REGION Network 343
   RUNG wire#powerrail
      Contact( "EMS".Carrier[46].SDC_OUT.Faults.CarrierSpacingFault )
      Coil( "Carrier_46_Carrier_Spacing_Fault" )
   END_RUNG
   // the same network as SCL:
   "Carrier_46_Carrier_Spacing_Fault" := "EMS".Carrier[46].SDC_OUT.Faults.CarrierSpacingFault;
END_REGION

REGION Network 344
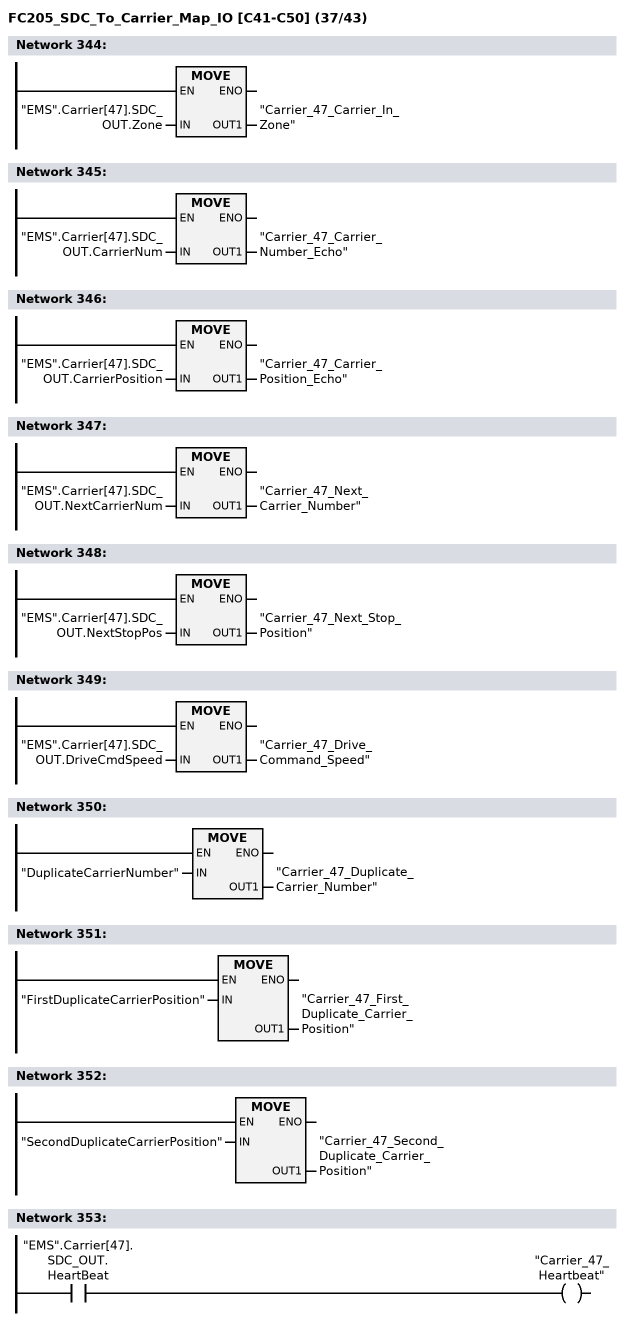
   RUNG wire#powerrail
      Move(in := "EMS".Carrier[47].SDC_OUT.Zone, out1 => "Carrier_47_Carrier_In_Zone")
   END_RUNG
   // the same network as SCL:
   "Carrier_47_Carrier_In_Zone" := "EMS".Carrier[47].SDC_OUT.Zone;
END_REGION

REGION Network 345
   RUNG wire#powerrail
      Move(in := "EMS".Carrier[47].SDC_OUT.CarrierNum, out1 => "Carrier_47_Carrier_Number_Echo")
   END_RUNG
   // the same network as SCL:
   "Carrier_47_Carrier_Number_Echo" := "EMS".Carrier[47].SDC_OUT.CarrierNum;
END_REGION

REGION Network 346
   RUNG wire#powerrail
      Move(in := "EMS".Carrier[47].SDC_OUT.CarrierPosition, out1 => "Carrier_47_Carrier_Position_Echo")
   END_RUNG
   // the same network as SCL:
   "Carrier_47_Carrier_Position_Echo" := "EMS".Carrier[47].SDC_OUT.CarrierPosition;
END_REGION

REGION Network 347
   RUNG wire#powerrail
      Move(in := "EMS".Carrier[47].SDC_OUT.NextCarrierNum, out1 => "Carrier_47_Next_Carrier_Number")
   END_RUNG
   // the same network as SCL:
   "Carrier_47_Next_Carrier_Number" := "EMS".Carrier[47].SDC_OUT.NextCarrierNum;
END_REGION

REGION Network 348
   RUNG wire#powerrail
      Move(in := "EMS".Carrier[47].SDC_OUT.NextStopPos, out1 => "Carrier_47_Next_Stop_Position")
   END_RUNG
   // the same network as SCL:
   "Carrier_47_Next_Stop_Position" := "EMS".Carrier[47].SDC_OUT.NextStopPos;
END_REGION

REGION Network 349
   RUNG wire#powerrail
      Move(in := "EMS".Carrier[47].SDC_OUT.DriveCmdSpeed, out1 => "Carrier_47_Drive_Command_Speed")
   END_RUNG
   // the same network as SCL:
   "Carrier_47_Drive_Command_Speed" := "EMS".Carrier[47].SDC_OUT.DriveCmdSpeed;
END_REGION

REGION Network 350
   RUNG wire#powerrail
      Move(in := "DuplicateCarrierNumber", out1 => "Carrier_47_Duplicate_Carrier_Number")
   END_RUNG
   // the same network as SCL:
   "Carrier_47_Duplicate_Carrier_Number" := "DuplicateCarrierNumber";
END_REGION

REGION Network 351
   RUNG wire#powerrail
      Move(in := "FirstDuplicateCarrierPosition", out1 => "Carrier_47_First_Duplicate_Carrier_Position")
   END_RUNG
   // the same network as SCL:
   "Carrier_47_First_Duplicate_Carrier_Position" := "FirstDuplicateCarrierPosition";
END_REGION

REGION Network 352
   RUNG wire#powerrail
      Move(in := "SecondDuplicateCarrierPosition", out1 => "Carrier_47_Second_Duplicate_Carrier_Position")
   END_RUNG
   // the same network as SCL:
   "Carrier_47_Second_Duplicate_Carrier_Position" := "SecondDuplicateCarrierPosition";
END_REGION

REGION Network 353
   RUNG wire#powerrail
      Contact( "EMS".Carrier[47].SDC_OUT.HeartBeat )
      Coil( "Carrier_47_Heartbeat" )
   END_RUNG
   // the same network as SCL:
   "Carrier_47_Heartbeat" := "EMS".Carrier[47].SDC_OUT.HeartBeat;
END_REGION

REGION Network 354
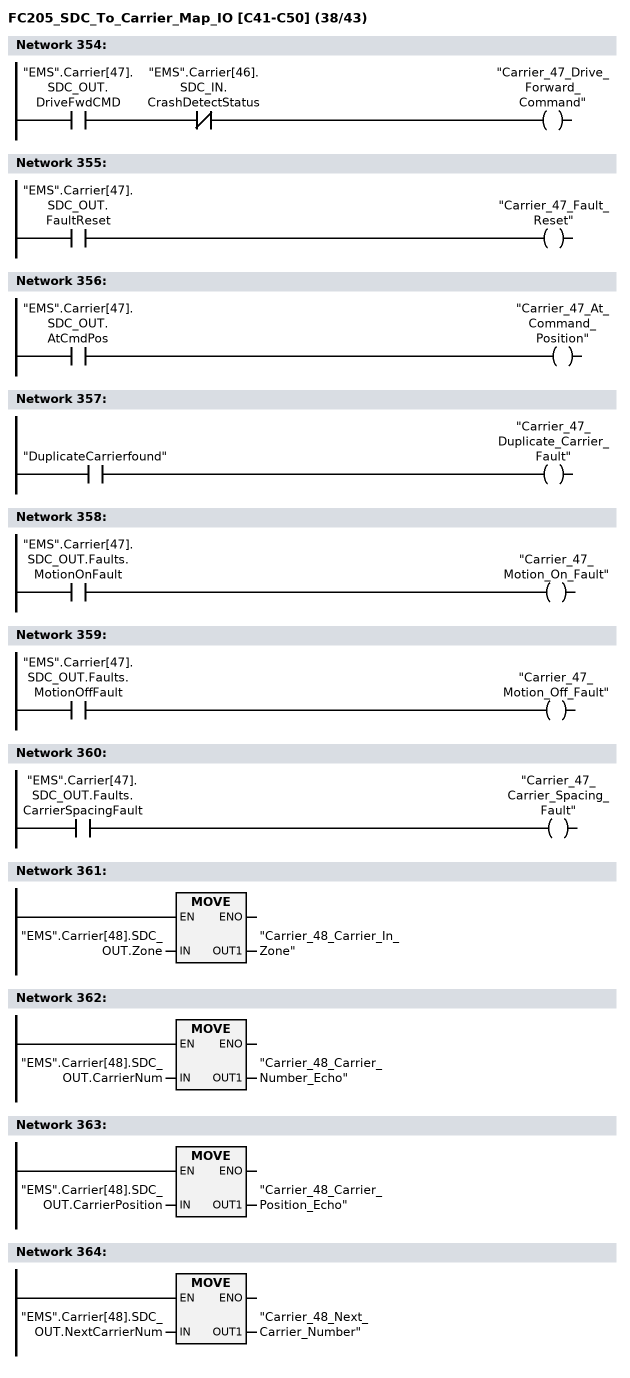
   RUNG wire#powerrail
      Contact( "EMS".Carrier[47].SDC_OUT.DriveFwdCMD )
      I_Contact( "EMS".Carrier[46].SDC_IN.CrashDetectStatus )
      Coil( "Carrier_47_Drive_Forward_Command" )
   END_RUNG
   // the same network as SCL:
   "Carrier_47_Drive_Forward_Command" := "EMS".Carrier[47].SDC_OUT.DriveFwdCMD AND NOT "EMS".Carrier[46].SDC_IN.CrashDetectStatus;
END_REGION

REGION Network 355
   RUNG wire#powerrail
      Contact( "EMS".Carrier[47].SDC_OUT.FaultReset )
      Coil( "Carrier_47_Fault_Reset" )
   END_RUNG
   // the same network as SCL:
   "Carrier_47_Fault_Reset" := "EMS".Carrier[47].SDC_OUT.FaultReset;
END_REGION

REGION Network 356
   RUNG wire#powerrail
      Contact( "EMS".Carrier[47].SDC_OUT.AtCmdPos )
      Coil( "Carrier_47_At_Command_Position" )
   END_RUNG
   // the same network as SCL:
   "Carrier_47_At_Command_Position" := "EMS".Carrier[47].SDC_OUT.AtCmdPos;
END_REGION

REGION Network 357
   RUNG wire#powerrail
      Contact( "DuplicateCarrierfound" )
      Coil( "Carrier_47_Duplicate_Carrier_Fault" )
   END_RUNG
   // the same network as SCL:
   "Carrier_47_Duplicate_Carrier_Fault" := "DuplicateCarrierfound";
END_REGION

REGION Network 358
   RUNG wire#powerrail
      Contact( "EMS".Carrier[47].SDC_OUT.Faults.MotionOnFault )
      Coil( "Carrier_47_Motion_On_Fault" )
   END_RUNG
   // the same network as SCL:
   "Carrier_47_Motion_On_Fault" := "EMS".Carrier[47].SDC_OUT.Faults.MotionOnFault;
END_REGION

REGION Network 359
   RUNG wire#powerrail
      Contact( "EMS".Carrier[47].SDC_OUT.Faults.MotionOffFault )
      Coil( "Carrier_47_Motion_Off_Fault" )
   END_RUNG
   // the same network as SCL:
   "Carrier_47_Motion_Off_Fault" := "EMS".Carrier[47].SDC_OUT.Faults.MotionOffFault;
END_REGION

REGION Network 360
   RUNG wire#powerrail
      Contact( "EMS".Carrier[47].SDC_OUT.Faults.CarrierSpacingFault )
      Coil( "Carrier_47_Carrier_Spacing_Fault" )
   END_RUNG
   // the same network as SCL:
   "Carrier_47_Carrier_Spacing_Fault" := "EMS".Carrier[47].SDC_OUT.Faults.CarrierSpacingFault;
END_REGION

REGION Network 361
   RUNG wire#powerrail
      Move(in := "EMS".Carrier[48].SDC_OUT.Zone, out1 => "Carrier_48_Carrier_In_Zone")
   END_RUNG
   // the same network as SCL:
   "Carrier_48_Carrier_In_Zone" := "EMS".Carrier[48].SDC_OUT.Zone;
END_REGION

REGION Network 362
   RUNG wire#powerrail
      Move(in := "EMS".Carrier[48].SDC_OUT.CarrierNum, out1 => "Carrier_48_Carrier_Number_Echo")
   END_RUNG
   // the same network as SCL:
   "Carrier_48_Carrier_Number_Echo" := "EMS".Carrier[48].SDC_OUT.CarrierNum;
END_REGION

REGION Network 363
   RUNG wire#powerrail
      Move(in := "EMS".Carrier[48].SDC_OUT.CarrierPosition, out1 => "Carrier_48_Carrier_Position_Echo")
   END_RUNG
   // the same network as SCL:
   "Carrier_48_Carrier_Position_Echo" := "EMS".Carrier[48].SDC_OUT.CarrierPosition;
END_REGION

REGION Network 364
   RUNG wire#powerrail
      Move(in := "EMS".Carrier[48].SDC_OUT.NextCarrierNum, out1 => "Carrier_48_Next_Carrier_Number")
   END_RUNG
   // the same network as SCL:
   "Carrier_48_Next_Carrier_Number" := "EMS".Carrier[48].SDC_OUT.NextCarrierNum;
END_REGION

REGION Network 365
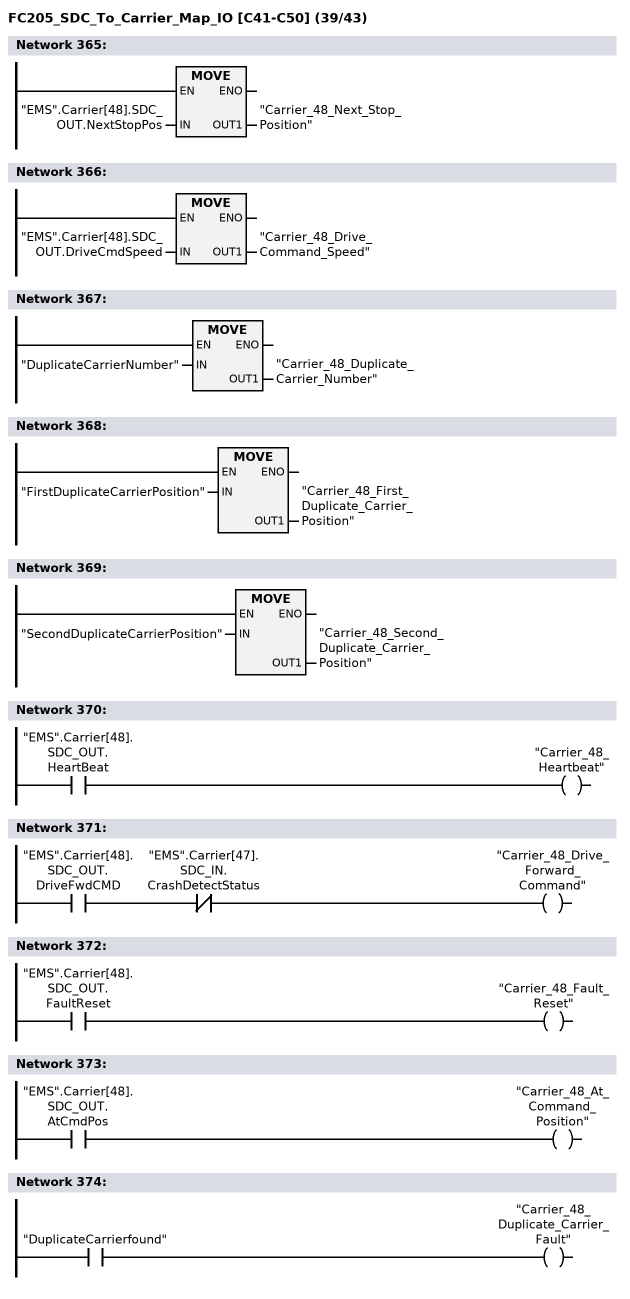
   RUNG wire#powerrail
      Move(in := "EMS".Carrier[48].SDC_OUT.NextStopPos, out1 => "Carrier_48_Next_Stop_Position")
   END_RUNG
   // the same network as SCL:
   "Carrier_48_Next_Stop_Position" := "EMS".Carrier[48].SDC_OUT.NextStopPos;
END_REGION

REGION Network 366
   RUNG wire#powerrail
      Move(in := "EMS".Carrier[48].SDC_OUT.DriveCmdSpeed, out1 => "Carrier_48_Drive_Command_Speed")
   END_RUNG
   // the same network as SCL:
   "Carrier_48_Drive_Command_Speed" := "EMS".Carrier[48].SDC_OUT.DriveCmdSpeed;
END_REGION

REGION Network 367
   RUNG wire#powerrail
      Move(in := "DuplicateCarrierNumber", out1 => "Carrier_48_Duplicate_Carrier_Number")
   END_RUNG
   // the same network as SCL:
   "Carrier_48_Duplicate_Carrier_Number" := "DuplicateCarrierNumber";
END_REGION

REGION Network 368
   RUNG wire#powerrail
      Move(in := "FirstDuplicateCarrierPosition", out1 => "Carrier_48_First_Duplicate_Carrier_Position")
   END_RUNG
   // the same network as SCL:
   "Carrier_48_First_Duplicate_Carrier_Position" := "FirstDuplicateCarrierPosition";
END_REGION

REGION Network 369
   RUNG wire#powerrail
      Move(in := "SecondDuplicateCarrierPosition", out1 => "Carrier_48_Second_Duplicate_Carrier_Position")
   END_RUNG
   // the same network as SCL:
   "Carrier_48_Second_Duplicate_Carrier_Position" := "SecondDuplicateCarrierPosition";
END_REGION

REGION Network 370
   RUNG wire#powerrail
      Contact( "EMS".Carrier[48].SDC_OUT.HeartBeat )
      Coil( "Carrier_48_Heartbeat" )
   END_RUNG
   // the same network as SCL:
   "Carrier_48_Heartbeat" := "EMS".Carrier[48].SDC_OUT.HeartBeat;
END_REGION

REGION Network 371
   RUNG wire#powerrail
      Contact( "EMS".Carrier[48].SDC_OUT.DriveFwdCMD )
      I_Contact( "EMS".Carrier[47].SDC_IN.CrashDetectStatus )
      Coil( "Carrier_48_Drive_Forward_Command" )
   END_RUNG
   // the same network as SCL:
   "Carrier_48_Drive_Forward_Command" := "EMS".Carrier[48].SDC_OUT.DriveFwdCMD AND NOT "EMS".Carrier[47].SDC_IN.CrashDetectStatus;
END_REGION

REGION Network 372
   RUNG wire#powerrail
      Contact( "EMS".Carrier[48].SDC_OUT.FaultReset )
      Coil( "Carrier_48_Fault_Reset" )
   END_RUNG
   // the same network as SCL:
   "Carrier_48_Fault_Reset" := "EMS".Carrier[48].SDC_OUT.FaultReset;
END_REGION

REGION Network 373
   RUNG wire#powerrail
      Contact( "EMS".Carrier[48].SDC_OUT.AtCmdPos )
      Coil( "Carrier_48_At_Command_Position" )
   END_RUNG
   // the same network as SCL:
   "Carrier_48_At_Command_Position" := "EMS".Carrier[48].SDC_OUT.AtCmdPos;
END_REGION

REGION Network 374
   RUNG wire#powerrail
      Contact( "DuplicateCarrierfound" )
      Coil( "Carrier_48_Duplicate_Carrier_Fault" )
   END_RUNG
   // the same network as SCL:
   "Carrier_48_Duplicate_Carrier_Fault" := "DuplicateCarrierfound";
END_REGION

REGION Network 375
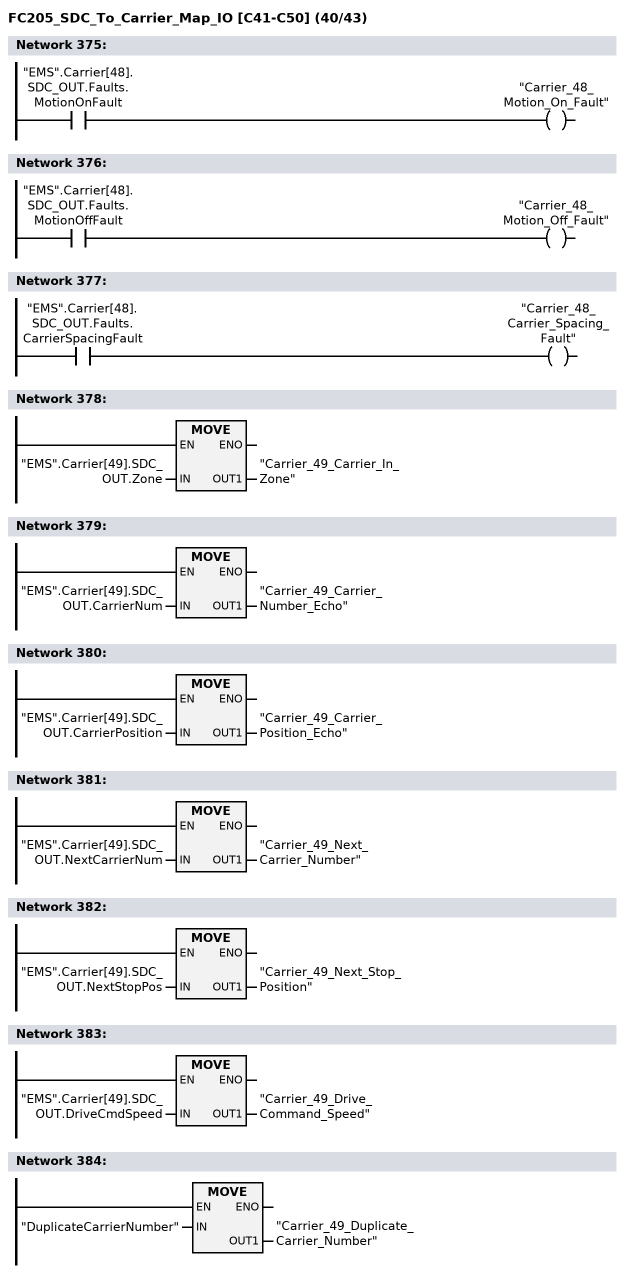
   RUNG wire#powerrail
      Contact( "EMS".Carrier[48].SDC_OUT.Faults.MotionOnFault )
      Coil( "Carrier_48_Motion_On_Fault" )
   END_RUNG
   // the same network as SCL:
   "Carrier_48_Motion_On_Fault" := "EMS".Carrier[48].SDC_OUT.Faults.MotionOnFault;
END_REGION

REGION Network 376
   RUNG wire#powerrail
      Contact( "EMS".Carrier[48].SDC_OUT.Faults.MotionOffFault )
      Coil( "Carrier_48_Motion_Off_Fault" )
   END_RUNG
   // the same network as SCL:
   "Carrier_48_Motion_Off_Fault" := "EMS".Carrier[48].SDC_OUT.Faults.MotionOffFault;
END_REGION

REGION Network 377
   RUNG wire#powerrail
      Contact( "EMS".Carrier[48].SDC_OUT.Faults.CarrierSpacingFault )
      Coil( "Carrier_48_Carrier_Spacing_Fault" )
   END_RUNG
   // the same network as SCL:
   "Carrier_48_Carrier_Spacing_Fault" := "EMS".Carrier[48].SDC_OUT.Faults.CarrierSpacingFault;
END_REGION

REGION Network 378
   RUNG wire#powerrail
      Move(in := "EMS".Carrier[49].SDC_OUT.Zone, out1 => "Carrier_49_Carrier_In_Zone")
   END_RUNG
   // the same network as SCL:
   "Carrier_49_Carrier_In_Zone" := "EMS".Carrier[49].SDC_OUT.Zone;
END_REGION

REGION Network 379
   RUNG wire#powerrail
      Move(in := "EMS".Carrier[49].SDC_OUT.CarrierNum, out1 => "Carrier_49_Carrier_Number_Echo")
   END_RUNG
   // the same network as SCL:
   "Carrier_49_Carrier_Number_Echo" := "EMS".Carrier[49].SDC_OUT.CarrierNum;
END_REGION

REGION Network 380
   RUNG wire#powerrail
      Move(in := "EMS".Carrier[49].SDC_OUT.CarrierPosition, out1 => "Carrier_49_Carrier_Position_Echo")
   END_RUNG
   // the same network as SCL:
   "Carrier_49_Carrier_Position_Echo" := "EMS".Carrier[49].SDC_OUT.CarrierPosition;
END_REGION

REGION Network 381
   RUNG wire#powerrail
      Move(in := "EMS".Carrier[49].SDC_OUT.NextCarrierNum, out1 => "Carrier_49_Next_Carrier_Number")
   END_RUNG
   // the same network as SCL:
   "Carrier_49_Next_Carrier_Number" := "EMS".Carrier[49].SDC_OUT.NextCarrierNum;
END_REGION

REGION Network 382
   RUNG wire#powerrail
      Move(in := "EMS".Carrier[49].SDC_OUT.NextStopPos, out1 => "Carrier_49_Next_Stop_Position")
   END_RUNG
   // the same network as SCL:
   "Carrier_49_Next_Stop_Position" := "EMS".Carrier[49].SDC_OUT.NextStopPos;
END_REGION

REGION Network 383
   RUNG wire#powerrail
      Move(in := "EMS".Carrier[49].SDC_OUT.DriveCmdSpeed, out1 => "Carrier_49_Drive_Command_Speed")
   END_RUNG
   // the same network as SCL:
   "Carrier_49_Drive_Command_Speed" := "EMS".Carrier[49].SDC_OUT.DriveCmdSpeed;
END_REGION

REGION Network 384
   RUNG wire#powerrail
      Move(in := "DuplicateCarrierNumber", out1 => "Carrier_49_Duplicate_Carrier_Number")
   END_RUNG
   // the same network as SCL:
   "Carrier_49_Duplicate_Carrier_Number" := "DuplicateCarrierNumber";
END_REGION

REGION Network 385
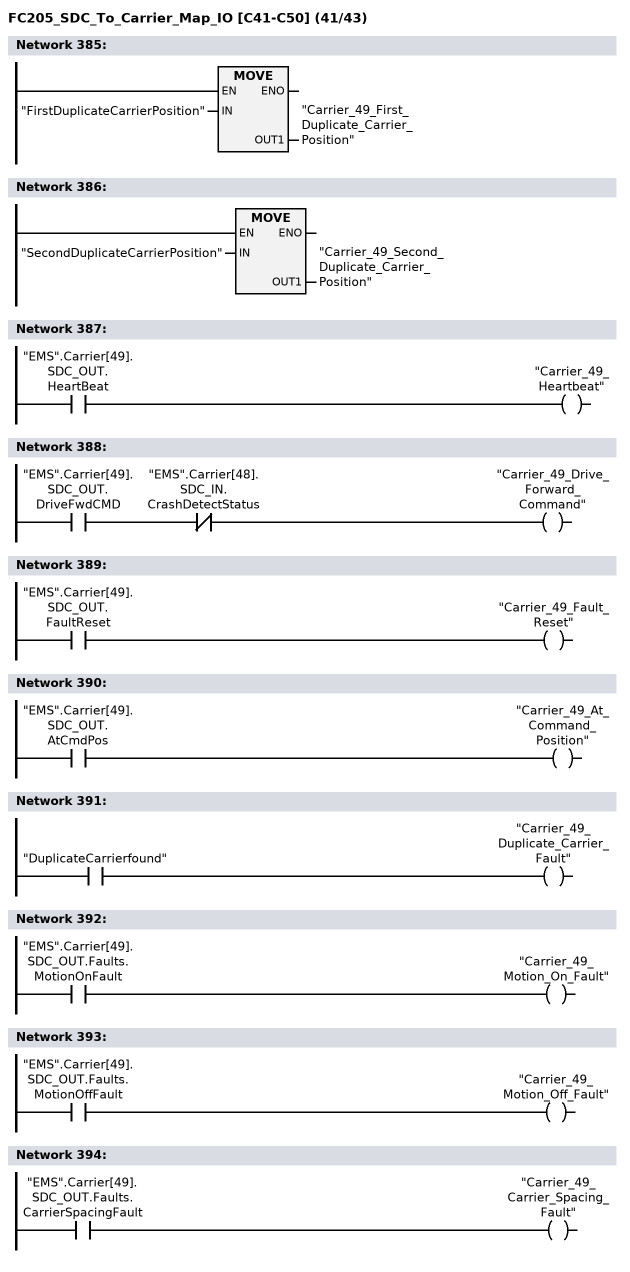
   RUNG wire#powerrail
      Move(in := "FirstDuplicateCarrierPosition", out1 => "Carrier_49_First_Duplicate_Carrier_Position")
   END_RUNG
   // the same network as SCL:
   "Carrier_49_First_Duplicate_Carrier_Position" := "FirstDuplicateCarrierPosition";
END_REGION

REGION Network 386
   RUNG wire#powerrail
      Move(in := "SecondDuplicateCarrierPosition", out1 => "Carrier_49_Second_Duplicate_Carrier_Position")
   END_RUNG
   // the same network as SCL:
   "Carrier_49_Second_Duplicate_Carrier_Position" := "SecondDuplicateCarrierPosition";
END_REGION

REGION Network 387
   RUNG wire#powerrail
      Contact( "EMS".Carrier[49].SDC_OUT.HeartBeat )
      Coil( "Carrier_49_Heartbeat" )
   END_RUNG
   // the same network as SCL:
   "Carrier_49_Heartbeat" := "EMS".Carrier[49].SDC_OUT.HeartBeat;
END_REGION

REGION Network 388
   RUNG wire#powerrail
      Contact( "EMS".Carrier[49].SDC_OUT.DriveFwdCMD )
      I_Contact( "EMS".Carrier[48].SDC_IN.CrashDetectStatus )
      Coil( "Carrier_49_Drive_Forward_Command" )
   END_RUNG
   // the same network as SCL:
   "Carrier_49_Drive_Forward_Command" := "EMS".Carrier[49].SDC_OUT.DriveFwdCMD AND NOT "EMS".Carrier[48].SDC_IN.CrashDetectStatus;
END_REGION

REGION Network 389
   RUNG wire#powerrail
      Contact( "EMS".Carrier[49].SDC_OUT.FaultReset )
      Coil( "Carrier_49_Fault_Reset" )
   END_RUNG
   // the same network as SCL:
   "Carrier_49_Fault_Reset" := "EMS".Carrier[49].SDC_OUT.FaultReset;
END_REGION

REGION Network 390
   RUNG wire#powerrail
      Contact( "EMS".Carrier[49].SDC_OUT.AtCmdPos )
      Coil( "Carrier_49_At_Command_Position" )
   END_RUNG
   // the same network as SCL:
   "Carrier_49_At_Command_Position" := "EMS".Carrier[49].SDC_OUT.AtCmdPos;
END_REGION

REGION Network 391
   RUNG wire#powerrail
      Contact( "DuplicateCarrierfound" )
      Coil( "Carrier_49_Duplicate_Carrier_Fault" )
   END_RUNG
   // the same network as SCL:
   "Carrier_49_Duplicate_Carrier_Fault" := "DuplicateCarrierfound";
END_REGION

REGION Network 392
   RUNG wire#powerrail
      Contact( "EMS".Carrier[49].SDC_OUT.Faults.MotionOnFault )
      Coil( "Carrier_49_Motion_On_Fault" )
   END_RUNG
   // the same network as SCL:
   "Carrier_49_Motion_On_Fault" := "EMS".Carrier[49].SDC_OUT.Faults.MotionOnFault;
END_REGION

REGION Network 393
   RUNG wire#powerrail
      Contact( "EMS".Carrier[49].SDC_OUT.Faults.MotionOffFault )
      Coil( "Carrier_49_Motion_Off_Fault" )
   END_RUNG
   // the same network as SCL:
   "Carrier_49_Motion_Off_Fault" := "EMS".Carrier[49].SDC_OUT.Faults.MotionOffFault;
END_REGION

REGION Network 394
   RUNG wire#powerrail
      Contact( "EMS".Carrier[49].SDC_OUT.Faults.CarrierSpacingFault )
      Coil( "Carrier_49_Carrier_Spacing_Fault" )
   END_RUNG
   // the same network as SCL:
   "Carrier_49_Carrier_Spacing_Fault" := "EMS".Carrier[49].SDC_OUT.Faults.CarrierSpacingFault;
END_REGION

REGION Network 395
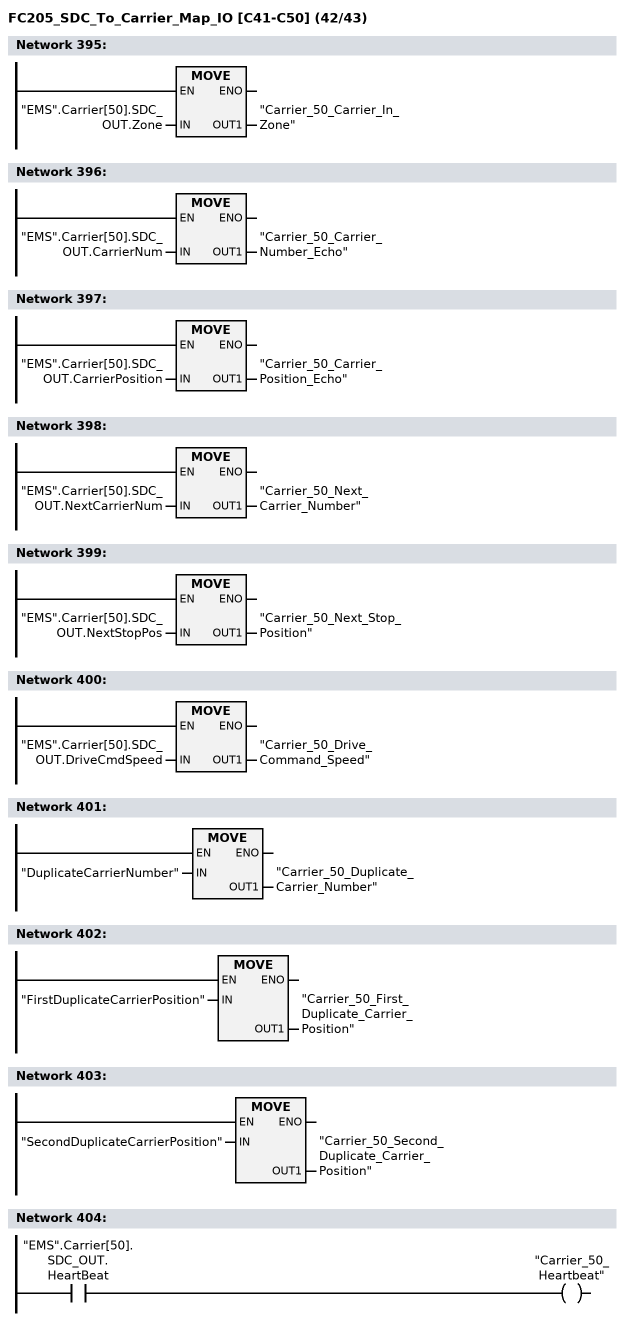
   RUNG wire#powerrail
      Move(in := "EMS".Carrier[50].SDC_OUT.Zone, out1 => "Carrier_50_Carrier_In_Zone")
   END_RUNG
   // the same network as SCL:
   "Carrier_50_Carrier_In_Zone" := "EMS".Carrier[50].SDC_OUT.Zone;
END_REGION

REGION Network 396
   RUNG wire#powerrail
      Move(in := "EMS".Carrier[50].SDC_OUT.CarrierNum, out1 => "Carrier_50_Carrier_Number_Echo")
   END_RUNG
   // the same network as SCL:
   "Carrier_50_Carrier_Number_Echo" := "EMS".Carrier[50].SDC_OUT.CarrierNum;
END_REGION

REGION Network 397
   RUNG wire#powerrail
      Move(in := "EMS".Carrier[50].SDC_OUT.CarrierPosition, out1 => "Carrier_50_Carrier_Position_Echo")
   END_RUNG
   // the same network as SCL:
   "Carrier_50_Carrier_Position_Echo" := "EMS".Carrier[50].SDC_OUT.CarrierPosition;
END_REGION

REGION Network 398
   RUNG wire#powerrail
      Move(in := "EMS".Carrier[50].SDC_OUT.NextCarrierNum, out1 => "Carrier_50_Next_Carrier_Number")
   END_RUNG
   // the same network as SCL:
   "Carrier_50_Next_Carrier_Number" := "EMS".Carrier[50].SDC_OUT.NextCarrierNum;
END_REGION

REGION Network 399
   RUNG wire#powerrail
      Move(in := "EMS".Carrier[50].SDC_OUT.NextStopPos, out1 => "Carrier_50_Next_Stop_Position")
   END_RUNG
   // the same network as SCL:
   "Carrier_50_Next_Stop_Position" := "EMS".Carrier[50].SDC_OUT.NextStopPos;
END_REGION

REGION Network 400
   RUNG wire#powerrail
      Move(in := "EMS".Carrier[50].SDC_OUT.DriveCmdSpeed, out1 => "Carrier_50_Drive_Command_Speed")
   END_RUNG
   // the same network as SCL:
   "Carrier_50_Drive_Command_Speed" := "EMS".Carrier[50].SDC_OUT.DriveCmdSpeed;
END_REGION

REGION Network 401
   RUNG wire#powerrail
      Move(in := "DuplicateCarrierNumber", out1 => "Carrier_50_Duplicate_Carrier_Number")
   END_RUNG
   // the same network as SCL:
   "Carrier_50_Duplicate_Carrier_Number" := "DuplicateCarrierNumber";
END_REGION

REGION Network 402
   RUNG wire#powerrail
      Move(in := "FirstDuplicateCarrierPosition", out1 => "Carrier_50_First_Duplicate_Carrier_Position")
   END_RUNG
   // the same network as SCL:
   "Carrier_50_First_Duplicate_Carrier_Position" := "FirstDuplicateCarrierPosition";
END_REGION

REGION Network 403
   RUNG wire#powerrail
      Move(in := "SecondDuplicateCarrierPosition", out1 => "Carrier_50_Second_Duplicate_Carrier_Position")
   END_RUNG
   // the same network as SCL:
   "Carrier_50_Second_Duplicate_Carrier_Position" := "SecondDuplicateCarrierPosition";
END_REGION

REGION Network 404
   RUNG wire#powerrail
      Contact( "EMS".Carrier[50].SDC_OUT.HeartBeat )
      Coil( "Carrier_50_Heartbeat" )
   END_RUNG
   // the same network as SCL:
   "Carrier_50_Heartbeat" := "EMS".Carrier[50].SDC_OUT.HeartBeat;
END_REGION

REGION Network 405
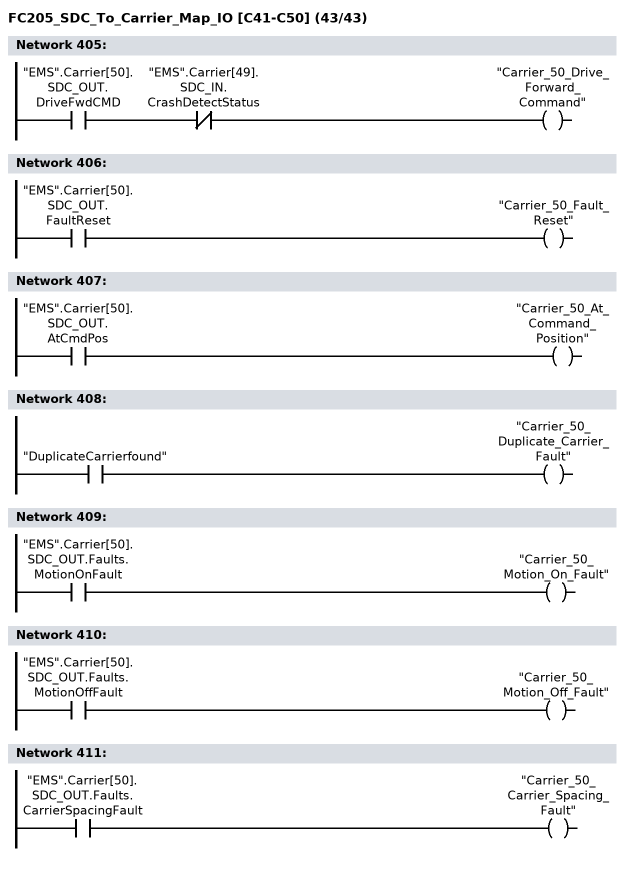
   RUNG wire#powerrail
      Contact( "EMS".Carrier[50].SDC_OUT.DriveFwdCMD )
      I_Contact( "EMS".Carrier[49].SDC_IN.CrashDetectStatus )
      Coil( "Carrier_50_Drive_Forward_Command" )
   END_RUNG
   // the same network as SCL:
   "Carrier_50_Drive_Forward_Command" := "EMS".Carrier[50].SDC_OUT.DriveFwdCMD AND NOT "EMS".Carrier[49].SDC_IN.CrashDetectStatus;
END_REGION

REGION Network 406
   RUNG wire#powerrail
      Contact( "EMS".Carrier[50].SDC_OUT.FaultReset )
      Coil( "Carrier_50_Fault_Reset" )
   END_RUNG
   // the same network as SCL:
   "Carrier_50_Fault_Reset" := "EMS".Carrier[50].SDC_OUT.FaultReset;
END_REGION

REGION Network 407
   RUNG wire#powerrail
      Contact( "EMS".Carrier[50].SDC_OUT.AtCmdPos )
      Coil( "Carrier_50_At_Command_Position" )
   END_RUNG
   // the same network as SCL:
   "Carrier_50_At_Command_Position" := "EMS".Carrier[50].SDC_OUT.AtCmdPos;
END_REGION

REGION Network 408
   RUNG wire#powerrail
      Contact( "DuplicateCarrierfound" )
      Coil( "Carrier_50_Duplicate_Carrier_Fault" )
   END_RUNG
   // the same network as SCL:
   "Carrier_50_Duplicate_Carrier_Fault" := "DuplicateCarrierfound";
END_REGION

REGION Network 409
   RUNG wire#powerrail
      Contact( "EMS".Carrier[50].SDC_OUT.Faults.MotionOnFault )
      Coil( "Carrier_50_Motion_On_Fault" )
   END_RUNG
   // the same network as SCL:
   "Carrier_50_Motion_On_Fault" := "EMS".Carrier[50].SDC_OUT.Faults.MotionOnFault;
END_REGION

REGION Network 410
   RUNG wire#powerrail
      Contact( "EMS".Carrier[50].SDC_OUT.Faults.MotionOffFault )
      Coil( "Carrier_50_Motion_Off_Fault" )
   END_RUNG
   // the same network as SCL:
   "Carrier_50_Motion_Off_Fault" := "EMS".Carrier[50].SDC_OUT.Faults.MotionOffFault;
END_REGION

REGION Network 411
   RUNG wire#powerrail
      Contact( "EMS".Carrier[50].SDC_OUT.Faults.CarrierSpacingFault )
      Coil( "Carrier_50_Carrier_Spacing_Fault" )
   END_RUNG
   // the same network as SCL:
   "Carrier_50_Carrier_Spacing_Fault" := "EMS".Carrier[50].SDC_OUT.Faults.CarrierSpacingFault;
END_REGION
END_FUNCTION

FUNCTION "FC206_SDC_To_Carrier_Map_IO [C51-C60]" : Void   // FC206, LAD
{ S7_Optimized_Access := 'TRUE' }
VERSION : 0.1
BEGIN

REGION Network 1
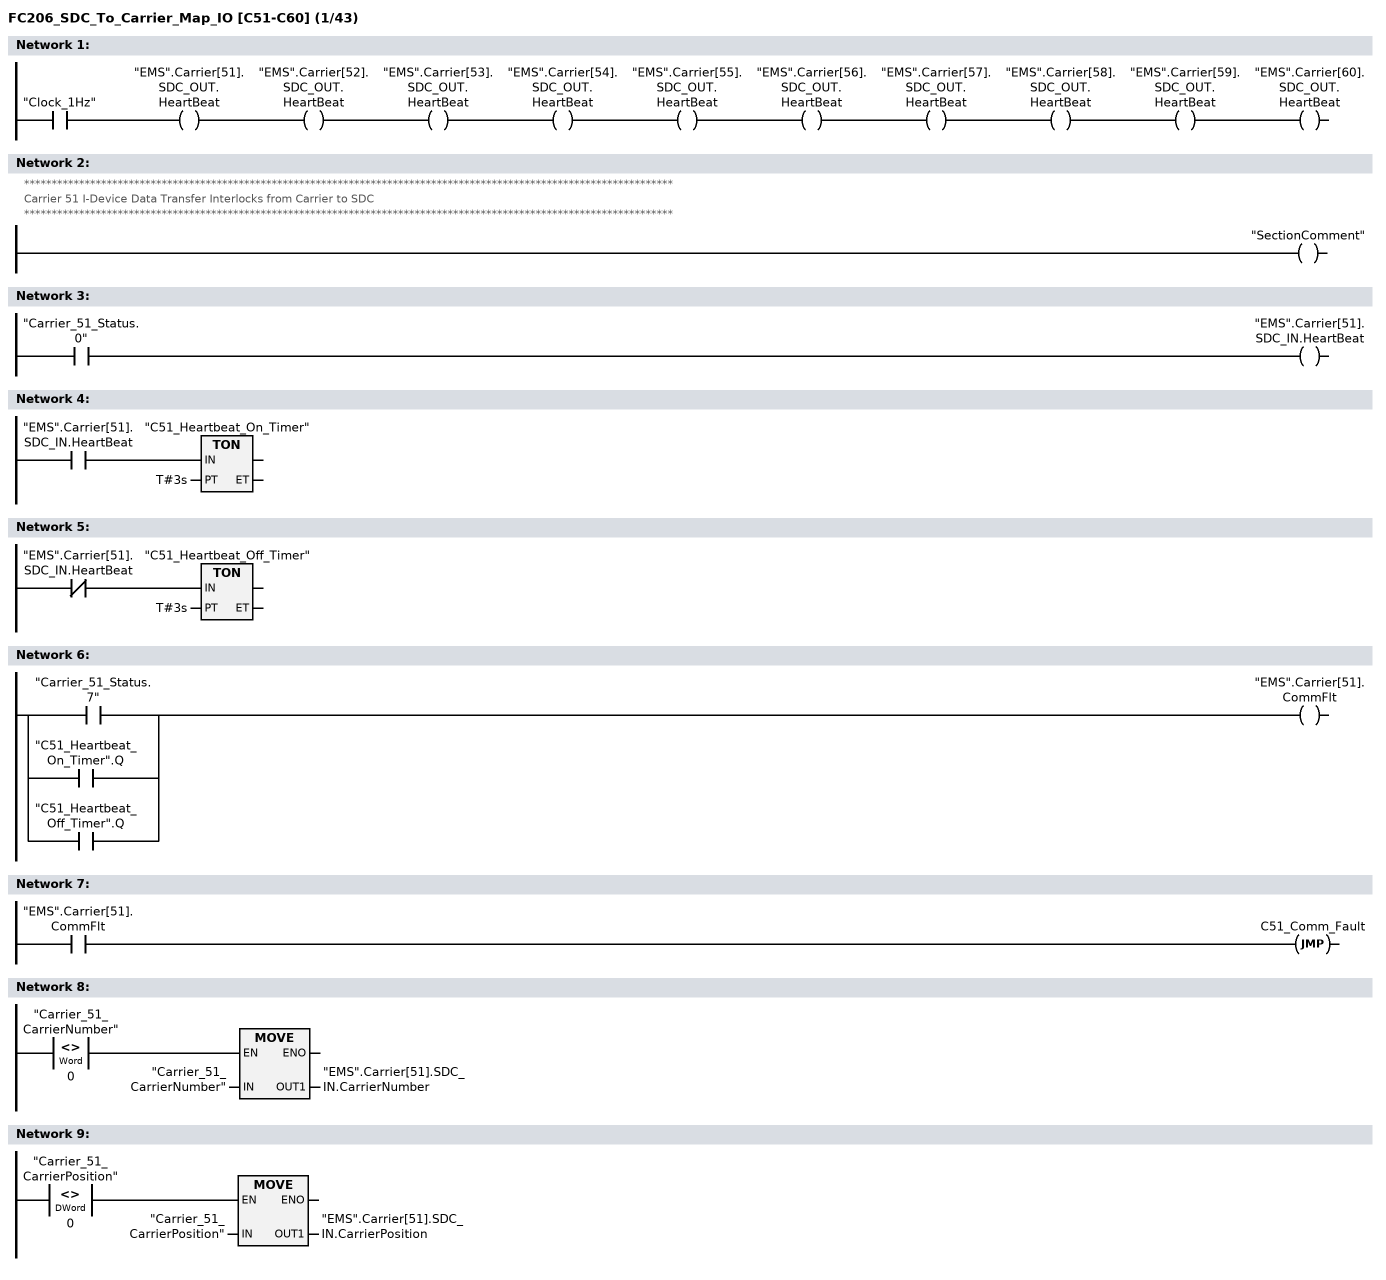
   RUNG wire#powerrail
      Contact( "Clock_1Hz" )
      Coil( "EMS".Carrier[51].SDC_OUT.HeartBeat )
      Coil( "EMS".Carrier[52].SDC_OUT.HeartBeat )
      Coil( "EMS".Carrier[53].SDC_OUT.HeartBeat )
      Coil( "EMS".Carrier[54].SDC_OUT.HeartBeat )
      Coil( "EMS".Carrier[55].SDC_OUT.HeartBeat )
      Coil( "EMS".Carrier[56].SDC_OUT.HeartBeat )
      Coil( "EMS".Carrier[57].SDC_OUT.HeartBeat )
      Coil( "EMS".Carrier[58].SDC_OUT.HeartBeat )
      Coil( "EMS".Carrier[59].SDC_OUT.HeartBeat )
      Coil( "EMS".Carrier[60].SDC_OUT.HeartBeat )
   END_RUNG
   // the same network as SCL:
   "EMS".Carrier[51].SDC_OUT.HeartBeat := "Clock_1Hz";
   "EMS".Carrier[52].SDC_OUT.HeartBeat := "Clock_1Hz";
   "EMS".Carrier[53].SDC_OUT.HeartBeat := "Clock_1Hz";
   "EMS".Carrier[54].SDC_OUT.HeartBeat := "Clock_1Hz";
   "EMS".Carrier[55].SDC_OUT.HeartBeat := "Clock_1Hz";
   "EMS".Carrier[56].SDC_OUT.HeartBeat := "Clock_1Hz";
   "EMS".Carrier[57].SDC_OUT.HeartBeat := "Clock_1Hz";
   "EMS".Carrier[58].SDC_OUT.HeartBeat := "Clock_1Hz";
   "EMS".Carrier[59].SDC_OUT.HeartBeat := "Clock_1Hz";
   "EMS".Carrier[60].SDC_OUT.HeartBeat := "Clock_1Hz";
END_REGION

REGION Network 2
   // **********************************************************************************************************************
   // 
   // Carrier 51 I-Device Data Transfer Interlocks from Carrier to SDC
   // 
   // **********************************************************************************************************************
   RUNG wire#powerrail
      Coil( "SectionComment" )
   END_RUNG
   // the same network as SCL:
   "SectionComment" := TRUE;
END_REGION

REGION Network 3
   RUNG wire#powerrail
      Contact( "Carrier_51_Status.0" )
      Coil( "EMS".Carrier[51].SDC_IN.HeartBeat )
   END_RUNG
   // the same network as SCL:
   "EMS".Carrier[51].SDC_IN.HeartBeat := "Carrier_51_Status.0";
END_REGION

REGION Network 4
   "C51_Heartbeat_On_Timer".TON(IN := "EMS".Carrier[51].SDC_IN.HeartBeat, PT := T#3s);
END_REGION

REGION Network 5
   "C51_Heartbeat_Off_Timer".TON(IN := NOT "EMS".Carrier[51].SDC_IN.HeartBeat, PT := T#3s);
END_REGION

REGION Network 6
   RUNG wire#powerrail
      Contact( "Carrier_51_Status.7" )
      wire#w1
      Coil( "EMS".Carrier[51].CommFlt )
   END_RUNG
   RUNG wire#powerrail
      Contact( "C51_Heartbeat_On_Timer".Q )
   END_RUNG wire#w1
   RUNG wire#powerrail
      Contact( "C51_Heartbeat_Off_Timer".Q )
   END_RUNG wire#w1
   // the same network as SCL:
   "EMS".Carrier[51].CommFlt := "Carrier_51_Status.7" OR "C51_Heartbeat_On_Timer".Q OR "C51_Heartbeat_Off_Timer".Q;
END_REGION

REGION Network 7
   RUNG wire#powerrail
      Contact( "EMS".Carrier[51].CommFlt )
      JumpCoil( C51_Comm_Fault )
   END_RUNG
   // the same network as SCL:
   IF "EMS".Carrier[51].CommFlt THEN GOTO C51_Comm_Fault; END_IF;
END_REGION

REGION Network 8
   RUNG wire#powerrail
      { S7_Templates := "SrcType := Word" } NE_Contact(in1 := "Carrier_51_CarrierNumber", in2 := 0)
      Move(in := "Carrier_51_CarrierNumber", out1 => "EMS".Carrier[51].SDC_IN.CarrierNumber)
   END_RUNG
   // the same network as SCL:
   IF "Carrier_51_CarrierNumber" <> 0 THEN
       "EMS".Carrier[51].SDC_IN.CarrierNumber := "Carrier_51_CarrierNumber";
   END_IF;
END_REGION

REGION Network 9
   RUNG wire#powerrail
      { S7_Templates := "SrcType := DWord" } NE_Contact(in1 := "Carrier_51_CarrierPosition", in2 := 0)
      Move(in := "Carrier_51_CarrierPosition", out1 => "EMS".Carrier[51].SDC_IN.CarrierPosition)
   END_RUNG
   // the same network as SCL:
   IF "Carrier_51_CarrierPosition" <> 0 THEN
       "EMS".Carrier[51].SDC_IN.CarrierPosition := "Carrier_51_CarrierPosition";
   END_IF;
END_REGION

REGION Network 10
